   "RIO3 Tanks Pressure Switch Hi Hi" : Bool = PLC "RIO3 Tanks Pressure Switch Hi Hi" AT %I33.1, 1 s
   "RIO3_SPR_DI_27_6" : Bool = PLC RIO3_SPR_DI_27_6 AT %I27.6, 1 s
   "RIO3_SPR_DI_27_7" : Bool = PLC RIO3_SPR_DI_27_7 AT %I27.7, 1 s
   "RIO3_SPR_DI_30_6" : Bool = PLC RIO3_SPR_DI_30_6 AT %I30.6, 1 s
   "RIO3_SPR_DI_30_7" : Bool = PLC RIO3_SPR_DI_30_7 AT %I30.7, 1 s
   "RIO3_SPR_DI_33_3" : Bool = PLC RIO3_SPR_DI_33_3 AT %I33.3, 1 s
   "RIO3_SPR_DI_33_4" : Bool = PLC RIO3_SPR_DI_33_4 AT %I33.4, 1 s
   "RIO3_SPR_DI_33_5" : Bool = PLC RIO3_SPR_DI_33_5 AT %I33.5, 1 s
   "RIO3_SPR_DI_33_6" : Bool = PLC RIO3_SPR_DI_33_6 AT %I33.6, 1 s
   "RIO3_SPR_DI_33_7" : Bool = PLC RIO3_SPR_DI_33_7 AT %I33.7, 1 s
   "RIO4 Tanks Pressure Switch Hi Hi" : Bool = PLC "RIO4 Tanks Pressure Switch Hi Hi" AT %I45.1, 1 s
   "RIO4_SPR_DI_139_6" : Bool = PLC RIO4_SPR_DI_139_6 AT %I39.6, 1 s
   "RIO4_SPR_DI_139_7" : Bool = PLC RIO4_SPR_DI_139_7 AT %I39.7, 1 s
   "RIO4_SPR_DI_142_6" : Bool = PLC RIO4_SPR_DI_142_6 AT %I42.6, 1 s
   "RIO4_SPR_DI_142_7" : Bool = PLC RIO4_SPR_DI_142_7 AT %I42.7, 1 s
   "RIO4_SPR_DI_145_3" : Bool = PLC RIO4_SPR_DI_145_3 AT %I45.3, 1 s
   "RIO4_SPR_DI_145_4" : Bool = PLC RIO4_SPR_DI_145_4 AT %I45.4, 1 s
   "RIO4_SPR_DI_145_5" : Bool = PLC RIO4_SPR_DI_145_5 AT %I45.5, 1 s
   "RIO4_SPR_DI_145_6" : Bool = PLC RIO4_SPR_DI_145_6 AT %I45.6, 1 s
   "RIO4_SPR_DI_145_7" : Bool = PLC RIO4_SPR_DI_145_7 AT %I45.7, 1 s
   "RIO5 Tanks Pressure Switch Hi Hi" : Bool = PLC "RIO5 Tanks Pressure Switch Hi Hi" AT %I57.1, 1 s
   "RIO5_SPR_DI_51_6" : Bool = PLC RIO5_SPR_DI_51_6 AT %I51.6, 1 s
   "RIO5_SPR_DI_51_7" : Bool = PLC RIO5_SPR_DI_51_7 AT %I51.7, 1 s
   "RIO5_SPR_DI_54_6" : Bool = PLC RIO5_SPR_DI_54_6 AT %I54.6, 1 s
   "RIO5_SPR_DI_54_7" : Bool = PLC RIO5_SPR_DI_54_7 AT %I54.7, 1 s
   "RIO5_SPR_DI_57_3" : Bool = PLC RIO5_SPR_DI_57_3 AT %I57.3, 1 s
   "RIO5_SPR_DI_57_4" : Bool = PLC RIO5_SPR_DI_57_4 AT %I57.4, 1 s
   "RIO5_SPR_DI_57_5" : Bool = PLC RIO5_SPR_DI_57_5 AT %I57.5, 1 s
   "RIO5_SPR_DI_57_6" : Bool = PLC RIO5_SPR_DI_57_6 AT %I57.6, 1 s
   "RIO5_SPR_DI_57_7" : Bool = PLC RIO5_SPR_DI_57_7 AT %I57.7, 1 s
   "RIO6 Tanks Pressure Switch Hi Hi" : Bool = PLC "RIO6 Tanks Pressure Switch Hi Hi" AT %I66.1, 1 s
   "RIO6_SPR_DI_60_6" : Bool = PLC RIO6_SPR_DI_60_6 AT %I60.6, 1 s
   "RIO6_SPR_DI_60_7" : Bool = PLC RIO6_SPR_DI_60_7 AT %I60.7, 1 s
   "RIO6_SPR_DI_63_6" : Bool = PLC RIO6_SPR_DI_63_6 AT %I63.6, 1 s
   "RIO6_SPR_DI_63_7" : Bool = PLC RIO6_SPR_DI_63_7 AT %I63.7, 1 s
   "RIO6_SPR_DI_66_3" : Bool = PLC RIO6_SPR_DI_66_3 AT %I66.3, 1 s
   "RIO6_SPR_DI_66_4" : Bool = PLC RIO6_SPR_DI_66_4 AT %I66.4, 1 s
   "RIO6_SPR_DI_66_5" : Bool = PLC RIO6_SPR_DI_66_5 AT %I66.5, 1 s
   "RIO6_SPR_DI_66_6" : Bool = PLC RIO6_SPR_DI_66_6 AT %I66.6, 1 s
   "RIO6_SPR_DI_66_7" : Bool = PLC RIO6_SPR_DI_66_7 AT %I66.7, 1 s
   "RIO7 Tank Pressure Switch Hi Hi" : Bool = PLC "RIO7 Tank Pressure Switch Hi Hi" AT %I78.1, 1 s
   "RIO7_SPR_DI_175_6" : Bool = PLC RIO7_SPR_DI_175_6 AT %I75.6, 1 s
   "RIO7_SPR_DI_175_7" : Bool = PLC RIO7_SPR_DI_175_7 AT %I75.7, 1 s
   "RIO7_SPR_DI_178_2" : Bool = PLC RIO7_SPR_DI_178_2 AT %I78.2, 1 s
   "RIO7_SPR_DI_178_3" : Bool = PLC RIO7_SPR_DI_178_3 AT %I78.3, 1 s
   "RIO7_SPR_DI_178_4" : Bool = PLC RIO7_SPR_DI_178_4 AT %I78.4, 1 s
   "RIO7_SPR_DI_178_5" : Bool = PLC RIO7_SPR_DI_178_5 AT %I78.5, 1 s
   "RIO7_SPR_DI_178_6" : Bool = PLC RIO7_SPR_DI_178_6 AT %I78.6, 1 s
   "RIO7_SPR_DI_178_7" : Bool = PLC RIO7_SPR_DI_178_7 AT %I78.7, 1 s
   "Safety System Interlock" : Bool = PLC "10_DI_Data".SFTY_SYS_IL AT %DB1.DBX0.0, 1 s
   "Sequence Times_DB_De-Ox SP Time" : Real = PLC "Sequence Times_DB"."De-Ox SP Time", 1 s
   "Sequence Times_DB_De-Ox Time" : Real = PLC "Sequence Times_DB"."De-Ox Time", 1 s
   "Sequence Times_DB_De-Ox Timer_Days Left" : DInt = PLC "Sequence Times_DB"."De-Ox Timer"."Days Left", 1 s
   "Sequence Times_DB_De-Ox Timer_Hours Left" : DInt = PLC "Sequence Times_DB"."De-Ox Timer"."Hours Left", 1 s
   "Sequence Times_DB_De-Ox Timer_Minutes Left" : DInt = PLC "Sequence Times_DB"."De-Ox Timer"."Minutes Left", 1 s
   "Sequence Times_DB_De-Ox Timer_PT_HOURS" : Real = PLC "Sequence Times_DB"."De-Ox Timer".PT_HOURS, 1 s
   "Sequence Times_DB_Dwell" : Real = PLC "Sequence Times_DB"."Dwell Time", 1 s
   "Sequence Times_DB_Dwell Timer_Days Left" : DInt = PLC "Sequence Times_DB"."Dwell Timer"."Days Left", 1 s
   "Sequence Times_DB_Dwell Timer_Hours Left" : DInt = PLC "Sequence Times_DB"."Dwell Timer"."Hours Left", 1 s
   "Sequence Times_DB_Dwell Timer_Minutes Left" : DInt = PLC "Sequence Times_DB"."Dwell Timer"."Minutes Left", 1 s
   "Sequence Times_DB_Dwell Timer_PT_HOURS" : Real = PLC "Sequence Times_DB"."Dwell Timer".PT_HOURS, 1 s
   "Sequence Times_DB_Jurney Time" : Real = PLC "Sequence Times_DB"."Jurney Time", 1 s
   "Sequence Times_DB_Jurney Time FB_Days Left" : Int = PLC "Sequence Times_DB"."Jurney Time FB"."Days Left", 1 s
   "Sequence Times_DB_Jurney Time FB_Hours Left" : Int = PLC "Sequence Times_DB"."Jurney Time FB"."Hours Left", 1 s
   "Sequence Times_DB_Jurney Time FB_PT_DAYS" : Real = PLC "Sequence Times_DB"."Jurney Time FB".PT_DAYS, 1 s
   "Sequence Times_DB_Jurney Timer_PT_DAYS" : Real = PLC "Sequence Times_DB"."Jurney Timer".PT_DAYS, 1 s
   "Sequence Times_DB_Jurney Timer_PT_HOURS" : Real = PLC "Sequence Times_DB"."Jurney Timer".PT_HOURS, 1 s
   "Sequence Times_DB_Jurney Timer_PT_MINUTES" : Real = PLC "Sequence Times_DB"."Jurney Timer".PT_MINUTES, 1 s
   "Sequence Times_DB_Post-Dwell" : Real = PLC "Sequence Times_DB"."Post-Dwell Time", 1 s
   "Sequence Times_DB_Post-Dwell Remaining_Days Left" : DInt = PLC "Sequence Times_DB"."Post-Dwell Timer"."Days Left", 1 s
   "Sequence Times_DB_Post-Dwell Remaining_Hours Left" : DInt = PLC "Sequence Times_DB"."Post-Dwell Timer"."Hours Left", 1 s
   "Sequence Times_DB_Post-Dwell Remaining_Minutes Left" : DInt = PLC "Sequence Times_DB"."Post-Dwell Timer"."Minutes Left", 1 s
   "Sequence Times_DB_Post-Dwell Remaining_PT_HOURS" : Real = PLC "Sequence Times_DB"."Post-Dwell Timer".PT_HOURS, 1 s
   "Sequence Times_DB_Pre-Dwell Time" : Real = PLC "Sequence Times_DB"."Pre-Dwell Time", 1 s
   "Sequence Times_DB_Pre-Dwell Timer_Days Left" : DInt = PLC "Sequence Times_DB"."Pre-Dwell Timer"."Days Left", 1 s
   "Sequence Times_DB_Pre-Dwell Timer_Hours Left" : DInt = PLC "Sequence Times_DB"."Pre-Dwell Timer"."Hours Left", 1 s
   "Sequence Times_DB_Pre-Dwell Timer_Minutes Left" : DInt = PLC "Sequence Times_DB"."Pre-Dwell Timer"."Minutes Left", 1 s
   "Sequence Times_DB_Pre-Dwell Timer_PT_DAYS" : Real = PLC "Sequence Times_DB"."Pre-Dwell Timer".PT_DAYS, 1 s
   "Sequence Times_DB_Pre-Dwell Timer_PT_HOURS" : Real = PLC "Sequence Times_DB"."Pre-Dwell Timer".PT_HOURS, 1 s
   "Sequence Times_DB_Pre-Dwell Timer_PT_MINUTES" : Real = PLC "Sequence Times_DB"."Pre-Dwell Timer".PT_MINUTES, 1 s
   "Sequence Times_DB_Re-Ox Time" : Real = PLC "Sequence Times_DB"."Re-Ox Time", 1 s
   "Sequence Times_DB_Re-Ox Timer_Days Left" : DInt = PLC "Sequence Times_DB"."Re-Ox Timer"."Days Left", 1 s
   "Sequence Times_DB_Re-Ox Timer_Hours Left" : DInt = PLC "Sequence Times_DB"."Re-Ox Timer"."Hours Left", 1 s
   "Sequence Times_DB_Re-Ox Timer_Minutes Left" : DInt = PLC "Sequence Times_DB"."Re-Ox Timer"."Minutes Left", 1 s
   "Sequence Times_DB_Re-Ox Timer_PT_HOURS" : Real = PLC "Sequence Times_DB"."Re-Ox Timer".PT_HOURS, 1 s
   "Sequence Times_DB_Treatment Timer_Days" : DInt = PLC "Sequence Times_DB"."Treatment Timer".Days, 1 s
   "Sequence Times_DB_Treatment Timer_Days Left" : DInt = PLC "Sequence Times_DB"."Treatment Timer"."Days Left", 1 s
   "Sequence Times_DB_Treatment Timer_Enable" : Bool = PLC "Sequence Times_DB"."Treatment Timer".Enable, 1 s
   "Sequence Times_DB_Treatment Timer_Hours" : DInt = PLC "Sequence Times_DB"."Treatment Timer".Hours, 1 s
   "Sequence Times_DB_Treatment Timer_Hours Left" : DInt = PLC "Sequence Times_DB"."Treatment Timer"."Hours Left", 1 s
   "Sequence Times_DB_Treatment Timer_Minutes" : DInt = PLC "Sequence Times_DB"."Treatment Timer".Minutes, 1 s
   "Sequence Times_DB_Treatment Timer_Minutes Left" : DInt = PLC "Sequence Times_DB"."Treatment Timer"."Minutes Left", 1 s
   "Shell Cooling Water Level Hi Hi Switch" : Bool = PLC "10 DI_DATA".LS001 AT %DB1.DBX0.0, 1 s
   "Shell CSW Temp Scaled" : Real = PLC "12_AI_Data".TIT315_SCALED AT %DB1.DBX0.0, 1 s
   "Shutdown" : Bool = PLC "14_DQ_Data".24PF2 AT %DB1.DBX0.0, 1 s
   "Shutdown Alarm" : Bool = PLC "14_DQ_Data".24K3 AT %DB1.DBX0.0, 1 s
   "Silence Buzzer" : Bool = PLC "80_From_HMI".SLNCE_BZR AT %DB1.DBX0.0, 1 s
   "Soot System Opacity" : Bool = PLC "10 DI_DATA".E700_OPACITY AT %DB1.DBX0.0, 1 s
   "Soot System Power Healthy" : Bool = PLC "10 DI_DATA".E700_PWR_OK AT %DB1.DBX0.0, 1 s
   "Spare Output BC Q1.2" : Bool = PLC "14_DQ_Data".R2_SPR_DQ_1_2 AT %DB1.DBX0.0, 1 s
   "Spare Output BC Q1.3" : Bool = PLC "14_DQ_Data".R2_SPR_DQ_1_3 AT %DB1.DBX0.0, 1 s
   "Spare Output BC Q1.4" : Bool = PLC "14_DQ_Data".R2_SPR_DQ_1_4 AT %DB1.DBX0.0, 1 s
   "Spare Output BC Q1.5" : Bool = PLC "14_DQ_Data".R2_SPR_DQ_1_5 AT %DB1.DBX0.0, 1 s
   "Spare Output BC Q1.6" : Bool = PLC "14_DQ_Data".R2_SPR_DQ_1_6 AT %DB1.DBX0.0, 1 s
   "Spare Output IGG Q0.7" : Bool = PLC "14_DQ_Data".R2_SPR_DQ_0_7 AT %DB1.DBX0.0, 1 s
   "Spare Output IGG Q1.0" : Bool = PLC "14_DQ_Data".R2_SPR_DQ_1_0 AT %DB1.DBX0.0, 1 s
   "Start IGG Flag" : Bool = PLC "80_From_HMI".RUN_IGG AT %DB1.DBX0.0, 1 s
   "Start Sequenc_DB_Post Purge Time Sec" : Int, internal
   "Tank 1P BWT Level High High Switch" : Bool = PLC "Tank 1P BWT Level High High Switch" AT %I9.2, 1 s
   "Tank 1P GTT Isolation Valve Feedback - Closed" : Bool = PLC "Tank 1P GTT Isolation Valve Feedback - Closed" AT %I3.1, 1 s
   "Tank 1P GTT Isolation Valve Feedback - Opened" : Bool = PLC "Tank 1P GTT Isolation Valve Feedback - Opened" AT %I3.0, 1 s
   "Tank 1P Tank Vent Valve 1 Feedback - Closed" : Bool = PLC "Tank 1P Tank Vent Valve 1 Feedback - Closed" AT %I3.3, 1 s
   "Tank 1P Tank Vent Valve 1 Feedback - Opened" : Bool = PLC "Tank 1P Tank Vent Valve 1 Feedback - Opened" AT %I3.2, 1 s
   "Tank 1P Tank Vent Valve 2 Feedback - Closed" : Bool = PLC "Tank 1P Tank Vent Valve 2 Feedback - Closed" AT %I3.5, 1 s
   "Tank 1P Tank Vent Valve 2 Feedback - Opened" : Bool = PLC "Tank 1P Tank Vent Valve 2 Feedback - Opened" AT %I3.4, 1 s
   "Tank 1S BWT Level High High Switch" : Bool = PLC "Tank 1S BWT Level High High Switch" AT %I9.3, 1 s
   "Tank 1S GTT Isolation Valve Feedback - Closed" : Bool = PLC "Tank 1S GTT Isolation Valve Feedback - Closed" AT %I6.1, 1 s
   "Tank 1S GTT Isolation Valve Feedback - Opened" : Bool = PLC "Tank 1S GTT Isolation Valve Feedback - Opened" AT %I6.0, 1 s
   "Tank 1S Tank Vent Valve 1 Feedback - Closed" : Bool = PLC "Tank 1S Tank Vent Valve 1 Feedback - Closed" AT %I6.3, 1 s
   "Tank 1S Tank Vent Valve 1 Feedback - Opened" : Bool = PLC "Tank 1S Tank Vent Valve 1 Feedback - Opened" AT %I6.2, 1 s
   "Tank 1S Tank Vent Valve 2 Feedback - Closed" : Bool = PLC "Tank 1S Tank Vent Valve 2 Feedback - Closed" AT %I6.5, 1 s
   "Tank 1S Tank Vent Valve 2 Feedback - Opened" : Bool = PLC "Tank 1S Tank Vent Valve 2 Feedback - Opened" AT %I6.4, 1 s
   "Tank 2P BWT Level High High Switch" : Bool = PLC "Tank 2P BWT Level High High Switch" AT %I21.0, 1 s
   "Tank 2P GTT Isolation Valve Feedback - Closed" : Bool = PLC "Tank 2P GTT Isolation Valve Feedback - Closed" AT %I15.1, 1 s
   "Tank 2P GTT Isolation Valve Feedback - Opened" : Bool = PLC "Tank 2P GTT Isolation Valve Feedback - Opened" AT %I15.0, 1 s
   "Tank 2P Tank Vent Valve 1 Feedback - Closed" : Bool = PLC "Tank 2P Tank Vent Valve 1 Feedback - Closed" AT %I15.3, 1 s
   "Tank 2P Tank Vent Valve 1 Feedback - Opened" : Bool = PLC "Tank 2P Tank Vent Valve 1 Feedback - Opened" AT %I15.2, 1 s
   "Tank 2P Tank Vent Valve 2 Feedback - Closed" : Bool = PLC "Tank 2P Tank Vent Valve 2 Feedback - Closed" AT %I15.5, 1 s
   "Tank 2P Tank Vent Valve 2 Feedback - Opened" : Bool = PLC "Tank 2P Tank Vent Valve 2 Feedback - Opened" AT %I15.4, 1 s
   "Tank 2S BWT Level High High Switch" : Bool = PLC "Tank 2S BWT Level High High Switch" AT %I21.2, 1 s
   "Tank 2S GTT Isolation Valve Feedback - Closed" : Bool = PLC "Tank 2S GTT Isolation Valve Feedback - Closed" AT %I18.1, 1 s
   "Tank 2S GTT Isolation Valve Feedback - Opened" : Bool = PLC "Tank 2S GTT Isolation Valve Feedback - Opened" AT %I18.0, 1 s
   "Tank 2S Tank Vent Valve 1 Feedback - Closed" : Bool = PLC "Tank 2S Tank Vent Valve 1 Feedback - Closed" AT %I18.3, 1 s
   "Tank 2S Tank Vent Valve 1 Feedback - Opened" : Bool = PLC "Tank 2S Tank Vent Valve 1 Feedback - Opened" AT %I18.2, 1 s
   "Tank 2S Tank Vent Valve 2 Feedback - Closed" : Bool = PLC "Tank 2S Tank Vent Valve 2 Feedback - Closed" AT %I18.5, 1 s
   "Tank 2S Tank Vent Valve 2 Feedback - Opened" : Bool = PLC "Tank 2S Tank Vent Valve 2 Feedback - Opened" AT %I18.4, 1 s
   "Tank 3P BWT Level High High Switch" : Bool = PLC "Tank 3P BWT Level High High Switch" AT %I33.0, 1 s
   "Tank 3P GTT Isolation Valve Feedback - Closed" : Bool = PLC "Tank 3P GTT Isolation Valve Feedback - Closed" AT %I27.1, 1 s
   "Tank 3P GTT Isolation Valve Feedback - Opened" : Bool = PLC "Tank 3P GTT Isolation Valve Feedback - Opened" AT %I27.0, 1 s
   "Tank 3P Tank Vent Valve 1 Feedback - Closed" : Bool = PLC "Tank 3P Tank Vent Valve 1 Feedback - Closed" AT %I27.3, 1 s
   "Tank 3P Tank Vent Valve 1 Feedback - Opened" : Bool = PLC "Tank 3P Tank Vent Valve 1 Feedback - Opened" AT %I27.2, 1 s
   "Tank 3P Tank Vent Valve 2 Feedback - Closed" : Bool = PLC "Tank 3P Tank Vent Valve 2 Feedback - Closed" AT %I27.5, 1 s
   "Tank 3P Tank Vent Valve 2 Feedback - Opened" : Bool = PLC "Tank 3P Tank Vent Valve 2 Feedback - Opened" AT %I27.4, 1 s
   "Tank 3S BWT Level High High Switch" : Bool = PLC "Tank 3S BWT Level High High Switch" AT %I33.2, 1 s
   "Tank 3S GTT Isolation Valve Feedback - Closed" : Bool = PLC "Tank 3S GTT Isolation Valve Feedback - Closed" AT %I30.1, 1 s
   "Tank 3S GTT Isolation Valve Feedback - Opened" : Bool = PLC "Tank 3S GTT Isolation Valve Feedback - Opened" AT %I30.0, 1 s
   "Tank 3S Tank Vent Valve 1 Feedback - Closed" : Bool = PLC "Tank 3S Tank Vent Valve 1 Feedback - Closed" AT %I30.3, 1 s
   "Tank 3S Tank Vent Valve 1 Feedback - Opened" : Bool = PLC "Tank 3S Tank Vent Valve 1 Feedback - Opened" AT %I30.2, 1 s
   "Tank 3S Tank Vent Valve 2 Feedback - Closed" : Bool = PLC "Tank 3S Tank Vent Valve 2 Feedback - Closed" AT %I30.5, 1 s
   "Tank 3S Tank Vent Valve 2 Feedback - Opened" : Bool = PLC "Tank 3S Tank Vent Valve 2 Feedback - Opened" AT %I30.4, 1 s
   "Tank 4P BWT Level High High Switch" : Bool = PLC "Tank 4P BWT Level High High Switch" AT %I45.0, 1 s
   "Tank 4P GTT Isolation Valve Feedback - Closed" : Bool = PLC "Tank 4P GTT Isolation Valve Feedback - Closed" AT %I39.1, 1 s
   "Tank 4P GTT Isolation Valve Feedback - Opened" : Bool = PLC "Tank 4P GTT Isolation Valve Feedback - Opened" AT %I39.0, 1 s
   "Tank 4P Tank Vent Valve 1 Feedback - Closed" : Bool = PLC "Tank 4P Tank Vent Valve 1 Feedback - Closed" AT %I39.3, 1 s
   "Tank 4P Tank Vent Valve 1 Feedback - Opened" : Bool = PLC "Tank 4P Tank Vent Valve 1 Feedback - Opened" AT %I39.2, 1 s
   "Tank 4P Tank Vent Valve 2 Feedback - Closed" : Bool = PLC "Tank 4P Tank Vent Valve 2 Feedback - Closed" AT %I39.5, 1 s
   "Tank 4P Tank Vent Valve 2 Feedback - Opened" : Bool = PLC "Tank 4P Tank Vent Valve 2 Feedback - Opened" AT %I39.4, 1 s
   "Tank 4S BWT Level High High Switch" : Bool = PLC "Tank 4S BWT Level High High Switch" AT %I45.2, 1 s
   "Tank 4S GTT Isolation Valve Feedback - Closed" : Bool = PLC "Tank 4S GTT Isolation Valve Feedback - Closed" AT %I42.1, 1 s
   "Tank 4S GTT Isolation Valve Feedback - Opened" : Bool = PLC "Tank 4S GTT Isolation Valve Feedback - Opened" AT %I42.0, 1 s
   "Tank 4S Tank Vent Valve 1 Feedback - Closed" : Bool = PLC "Tank 4S Tank Vent Valve 1 Feedback - Closed" AT %I42.3, 1 s
   "Tank 4S Tank Vent Valve 1 Feedback - Opened" : Bool = PLC "Tank 4S Tank Vent Valve 1 Feedback - Opened" AT %I42.2, 1 s
   "Tank 4S Tank Vent Valve 2 Feedback - Closed" : Bool = PLC "Tank 4S Tank Vent Valve 2 Feedback - Closed" AT %I42.5, 1 s
   "Tank 4S Tank Vent Valve 2 Feedback - Opened" : Bool = PLC "Tank 4S Tank Vent Valve 2 Feedback - Opened" AT %I42.4, 1 s
   "Tank 5P BWT Level High High Switch" : Bool = PLC "Tank 5P BWT Level High High Switch" AT %I57.0, 1 s
   "Tank 5P GTT Isolation Valve Feedback - Closed" : Bool = PLC "Tank 5P GTT Isolation Valve Feedback - Closed" AT %I51.1, 1 s
   "Tank 5P GTT Isolation Valve Feedback - Opened" : Bool = PLC "Tank 5P GTT Isolation Valve Feedback - Opened" AT %I51.0, 1 s
   "Tank 5P Tank Vent Valve 1 Feedback - Closed" : Bool = PLC "Tank 5P Tank Vent Valve 1 Feedback - Closed" AT %I51.3, 1 s
   "Tank 5P Tank Vent Valve 1 Feedback - Opened" : Bool = PLC "Tank 5P Tank Vent Valve 1 Feedback - Opened" AT %I51.2, 1 s
   "Tank 5P Tank Vent Valve 2 Feedback - Closed" : Bool = PLC "Tank 5P Tank Vent Valve 2 Feedback - Closed" AT %I51.5, 1 s
   "Tank 5P Tank Vent Valve 2 Feedback - Opened" : Bool = PLC "Tank 5P Tank Vent Valve 2 Feedback - Opened" AT %I51.4, 1 s
   "Tank 5S BWT Level High High Switch" : Bool = PLC "Tank 5S BWT Level High High Switch" AT %I57.2, 1 s
   "Tank 6P BWT Level High High Switch" : Bool = PLC "Tank 6P BWT Level High High Switch" AT %I66.0, 1 s
   "Tank 6S BWT Level High High Switch" : Bool = PLC "Tank 6S BWT Level High High Switch" AT %I66.2, 1 s
   "Test Pressure Valve Control" : Bool = PLC "14_DQ_Data".200CV127ControlOut AT %DB1.DBX0.0, 1 s
   "TIT406_ALM_ANALOG_DB74_HIGH LEVEL VALUE (H)" : Real = PLC TIT406_ALM_ANALOG_DB74."HIGH LEVEL VALUE (H)" AT %DB74.DBD30, 1 s
   "TIT406_ALM_ANALOG_DB74_LOW LEVEL VALUE (L)" : Real = PLC TIT406_ALM_ANALOG_DB74."LOW LEVEL VALUE (L)" AT %DB74.DBD26, 1 s
   "TIT406_ALM_ANALOG_DB74_VERY HIGH LEVEL VALUE (HH)" : Real = PLC TIT406_ALM_ANALOG_DB74."VERY HIGH LEVEL VALUE (HH)" AT %DB74.DBD34, 1 s
   "TIT406_ALM_ANALOG_DB74_VERY LOW LEVEL VALUE (LL)" : Real = PLC TIT406_ALM_ANALOG_DB74."VERY LOW LEVEL VALUE (LL)" AT %DB74.DBD22, 1 s
   "TIT408_ALM_ANALOG_DB75_HIGH LEVEL VALUE (H)" : Real = PLC TIT408_ALM_ANALOG_DB75."HIGH LEVEL VALUE (H)" AT %DB75.DBD30, 1 s
   "TIT408_ALM_ANALOG_DB75_LOW LEVEL VALUE (L)" : Real = PLC TIT408_ALM_ANALOG_DB75."LOW LEVEL VALUE (L)" AT %DB75.DBD26, 1 s
   "TIT408_ALM_ANALOG_DB75_VERY HIGH LEVEL VALUE (HH)" : Real = PLC TIT408_ALM_ANALOG_DB75."VERY HIGH LEVEL VALUE (HH)" AT %DB75.DBD34, 1 s
   "TIT408_ALM_ANALOG_DB75_VERY LOW LEVEL VALUE (LL)" : Real = PLC TIT408_ALM_ANALOG_DB75."VERY LOW LEVEL VALUE (LL)" AT %DB75.DBD22, 1 s
   "Treatment Runs Completed" : Bool = PLC "2102_TIME_CALCS_DB".POST_DWELL_TMR_DN AT %DB1.DBD0, 1 s
   "user_group" : Int, internal
   "Vent Valve Control HMI Position" : Real = PLC "16_AQ_Data".CV403_CNTRL AT %DB1.DBX0.0, 1 s
   "Vent Valve Position Control" : Real = PLC "12_AI_Data".CV403_SCALED AT %DB1.DBX0.0, 1 s
   "Voyage_TIME_exceded" : Bool = PLC "2102_TIME_CALCS_DB".Voyage_TIME_invalid AT %DB1.DBW0, 1 s
   "Warning Alarm" : Bool = PLC "14_DQ_Data".24PF3 AT %DB1.DBX0.0, 1 s
   "Sequence Times_DB_Continue" : Bool = PLC "Sequence Times_DB".Continue, 1 s
   "Recipe Tag" : Int AT %DB1.DBX0.0
   "Record Data Tag" : Int AT %DB1.DBX0.0
   "Data_From_WBT_Level_APT" : Real = PLC Data_From_WBT.Level_APT, 1 s
   "Data_From_WBT_Level_WBT_6P" : Real = PLC Data_From_WBT.Level_WBT_6P, 1 s
   "Data_From_WBT_Level_WBT_5P" : Real = PLC Data_From_WBT.Level_WBT_5P, 1 s
   "Data_From_WBT_Level_WBT_4P" : Real = PLC Data_From_WBT.Level_WBT_4P, 1 s
   "Data_From_WBT_Level_WBT_3P" : Real = PLC Data_From_WBT.Level_WBT_3P, 1 s
   "Data_From_WBT_Level_WBT_2P" : Real = PLC Data_From_WBT.Level_WBT_2P, 1 s
   "Data_From_WBT_Level_WBT_1P" : Real = PLC Data_From_WBT.Level_WBT_1P, 1 s
   "Data_From_WBT_Level_FPT" : Real = PLC Data_From_WBT.Level_FPT, 1 s
   "Data_From_WBT_Level_WBT_1S" : Real = PLC Data_From_WBT.Level_WBT_1S, 1 s
   "Data_From_WBT_Level_WBT_2S" : Real = PLC Data_From_WBT.Level_WBT_2S, 1 s
   "Data_From_WBT_Level_WBT_3S" : Real = PLC Data_From_WBT.Level_WBT_3S, 1 s
   "Data_From_WBT_Level_WBT_4S" : Real = PLC Data_From_WBT.Level_WBT_4S, 1 s
   "Data_From_WBT_Level_WBT_5S" : Real = PLC Data_From_WBT.Level_WBT_5S, 1 s
   "Data_From_WBT_Level_WBT_6S" : Real = PLC Data_From_WBT.Level_WBT_6S, 1 s
   "IN_Level_APT" : Int = PLC IN_Level_APT AT %IW1026, 1 s
   "Data_From_WBT_Level_APT m" : Real = PLC Data_From_WBT."Level_APT m", 1 s
   "Data_From_WBT_Level_WBT_6S m" : Real = PLC Data_From_WBT."Level_WBT_6S m", 1 s
   "Data_From_WBT_Level_WBT_5S m" : Real = PLC Data_From_WBT."Level_WBT_5S m", 1 s
   "Data_From_WBT_Level_WBT_4S m" : Real = PLC Data_From_WBT."Level_WBT_4S m", 1 s
   "Data_From_WBT_Level_WBT_3S m" : Real = PLC Data_From_WBT."Level_WBT_3S m", 1 s
   "Data_From_WBT_Level_WBT_2S m" : Real = PLC Data_From_WBT."Level_WBT_2S m", 1 s
   "Data_From_WBT_Level_WBT_1S m" : Real = PLC Data_From_WBT."Level_WBT_1S m", 1 s
   "Data_From_WBT_Level_FPT m" : Real = PLC Data_From_WBT."Level_FPT m", 1 s
   "Data_From_WBT_Level_WBT_1P m" : Real = PLC Data_From_WBT."Level_WBT_1P m", 1 s
   "Data_From_WBT_Level_WBT_2P m" : Real = PLC Data_From_WBT."Level_WBT_2P m", 1 s
   "Data_From_WBT_Level_WBT_3P m" : Real = PLC Data_From_WBT."Level_WBT_3P m", 1 s
   "Data_From_WBT_Level_WBT_4P m" : Real = PLC Data_From_WBT."Level_WBT_4P m", 1 s
   "Data_From_WBT_Level_WBT_5P m" : Real = PLC Data_From_WBT."Level_WBT_5P m", 1 s
   "Data_From_WBT_Level_WBT_6P m" : Real = PLC Data_From_WBT."Level_WBT_6P m", 1 s
   "Alarm beacon handling_DB_Warning" : Bool = PLC "Alarm beacon handling_DB".Warning, 1 s
   "Alarm beacon handling_DB_Alarm" : Bool = PLC "Alarm beacon handling_DB".Alarm, 1 s
   "63_Safety System Interlock_IDB_Lockout Healthy" : Bool = PLC "63_Safety System Interlock_IDB"."Lockout Healthy", 1 s
   "63_Safety System Interlock_IDB_Reset Lockout" : Bool = PLC "63_Safety System Interlock_IDB"."Reset Lockout", 1 s
   "IDB_E131_Functioning Hours_Service Time bit" : Bool = PLC "IDB_E131_Functioning Hours"."Service Time bit", 1 s
   "Operation hours E139_IDB_Service Time bit" : Bool = PLC "Operation hours E139_IDB"."Service Time bit", 1 s
   "E-400 Animation_DB_Animation" : Int = PLC "E-400 Animation_DB".Animation, 1 s
   "20_TANKS_IP_DATA_RIO_01_FIRST_TANK_TANK_ALARM" : Bool = PLC "20_TANKS_IP_DATA".RIO_01.FIRST_TANK.TANK_ALARM, 1 s
   "CSW_Animation_DB_Animation" : Int = PLC CSW_Animation_DB.Animation, 1 s
   "103_Main_Burner_DB_FLM_DET" : Bool = PLC "103_Main_Burner_DB".FLM_DET, 1 s
   "504_Tank Grouping_DB2020_Time Left Tank_Time Left d Tank 1" : DInt = PLC "504_Tank Grouping_DB2020"."Time Left Tank"."Time Left d Tank 1", 1 s
   "504_Tank Grouping_DB2020_Time Left Tank_Time Left d Tank 10" : DInt = PLC "504_Tank Grouping_DB2020"."Time Left Tank"."Time Left d Tank 10", 1 s
   "504_Tank Grouping_DB2020_Time Left Tank_Time Left d Tank 11" : DInt = PLC "504_Tank Grouping_DB2020"."Time Left Tank"."Time Left d Tank 11", 1 s
   "504_Tank Grouping_DB2020_Time Left Tank_Time Left d Tank 12" : DInt = PLC "504_Tank Grouping_DB2020"."Time Left Tank"."Time Left d Tank 12", 1 s
   "504_Tank Grouping_DB2020_Time Left Tank_Time Left d Tank 13" : DInt = PLC "504_Tank Grouping_DB2020"."Time Left Tank"."Time Left d Tank 13", 1 s
   "504_Tank Grouping_DB2020_Time Left Tank_Time Left d Tank 14" : DInt = PLC "504_Tank Grouping_DB2020"."Time Left Tank"."Time Left d Tank 14", 1 s
   "504_Tank Grouping_DB2020_Time Left Tank_Time Left d Tank 2" : DInt = PLC "504_Tank Grouping_DB2020"."Time Left Tank"."Time Left d Tank 2", 1 s
   "504_Tank Grouping_DB2020_Time Left Tank_Time Left d Tank 3" : DInt = PLC "504_Tank Grouping_DB2020"."Time Left Tank"."Time Left d Tank 3", 1 s
   "504_Tank Grouping_DB2020_Time Left Tank_Time Left d Tank 4" : DInt = PLC "504_Tank Grouping_DB2020"."Time Left Tank"."Time Left d Tank 4", 1 s
   "504_Tank Grouping_DB2020_Time Left Tank_Time Left d Tank 5" : DInt = PLC "504_Tank Grouping_DB2020"."Time Left Tank"."Time Left d Tank 5", 1 s
   "504_Tank Grouping_DB2020_Time Left Tank_Time Left d Tank 6" : DInt = PLC "504_Tank Grouping_DB2020"."Time Left Tank"."Time Left d Tank 6", 1 s
   "504_Tank Grouping_DB2020_Time Left Tank_Time Left d Tank 7" : DInt = PLC "504_Tank Grouping_DB2020"."Time Left Tank"."Time Left d Tank 7", 1 s
   "504_Tank Grouping_DB2020_Time Left Tank_Time Left d Tank 8" : DInt = PLC "504_Tank Grouping_DB2020"."Time Left Tank"."Time Left d Tank 8", 1 s
   "504_Tank Grouping_DB2020_Time Left Tank_Time Left d Tank 9" : DInt = PLC "504_Tank Grouping_DB2020"."Time Left Tank"."Time Left d Tank 9", 1 s
   "504_Tank Grouping_DB2020_Time Left Tank_Time Left h Tank 1" : DInt = PLC "504_Tank Grouping_DB2020"."Time Left Tank"."Time Left h Tank 1", 1 s
   "504_Tank Grouping_DB2020_Time Left Tank_Time Left h Tank 10" : DInt = PLC "504_Tank Grouping_DB2020"."Time Left Tank"."Time Left h Tank 10", 1 s
   "504_Tank Grouping_DB2020_Time Left Tank_Time Left h Tank 11" : DInt = PLC "504_Tank Grouping_DB2020"."Time Left Tank"."Time Left h Tank 11", 1 s
   "504_Tank Grouping_DB2020_Time Left Tank_Time Left h Tank 12" : DInt = PLC "504_Tank Grouping_DB2020"."Time Left Tank"."Time Left h Tank 12", 1 s
   "504_Tank Grouping_DB2020_Time Left Tank_Time Left h Tank 13" : DInt = PLC "504_Tank Grouping_DB2020"."Time Left Tank"."Time Left h Tank 13", 1 s
   "504_Tank Grouping_DB2020_Time Left Tank_Time Left h Tank 14" : DInt = PLC "504_Tank Grouping_DB2020"."Time Left Tank"."Time Left h Tank 14", 1 s
   "504_Tank Grouping_DB2020_Time Left Tank_Time Left h Tank 2" : DInt = PLC "504_Tank Grouping_DB2020"."Time Left Tank"."Time Left h Tank 2", 1 s
   "504_Tank Grouping_DB2020_Time Left Tank_Time Left h Tank 3" : DInt = PLC "504_Tank Grouping_DB2020"."Time Left Tank"."Time Left h Tank 3", 1 s
   "504_Tank Grouping_DB2020_Time Left Tank_Time Left h Tank 4" : DInt = PLC "504_Tank Grouping_DB2020"."Time Left Tank"."Time Left h Tank 4", 1 s
   "504_Tank Grouping_DB2020_Time Left Tank_Time Left h Tank 5" : DInt = PLC "504_Tank Grouping_DB2020"."Time Left Tank"."Time Left h Tank 5", 1 s
   "504_Tank Grouping_DB2020_Time Left Tank_Time Left h Tank 6" : DInt = PLC "504_Tank Grouping_DB2020"."Time Left Tank"."Time Left h Tank 6", 1 s
   "504_Tank Grouping_DB2020_Time Left Tank_Time Left h Tank 7" : DInt = PLC "504_Tank Grouping_DB2020"."Time Left Tank"."Time Left h Tank 7", 1 s
   "504_Tank Grouping_DB2020_Time Left Tank_Time Left h Tank 8" : DInt = PLC "504_Tank Grouping_DB2020"."Time Left Tank"."Time Left h Tank 8", 1 s
   "504_Tank Grouping_DB2020_Time Left Tank_Time Left h Tank 9" : DInt = PLC "504_Tank Grouping_DB2020"."Time Left Tank"."Time Left h Tank 9", 1 s
   "504_Tank Grouping_DB2020_Time Left Tank_Time Left m Tank 1" : DInt = PLC "504_Tank Grouping_DB2020"."Time Left Tank"."Time Left m Tank 1", 1 s
   "504_Tank Grouping_DB2020_Time Left Tank_Time Left m Tank 10" : DInt = PLC "504_Tank Grouping_DB2020"."Time Left Tank"."Time Left m Tank 10", 1 s
   "504_Tank Grouping_DB2020_Time Left Tank_Time Left m Tank 11" : DInt = PLC "504_Tank Grouping_DB2020"."Time Left Tank"."Time Left m Tank 11", 1 s
   "504_Tank Grouping_DB2020_Time Left Tank_Time Left m Tank 12" : DInt = PLC "504_Tank Grouping_DB2020"."Time Left Tank"."Time Left m Tank 12", 1 s
   "504_Tank Grouping_DB2020_Time Left Tank_Time Left m Tank 13" : DInt = PLC "504_Tank Grouping_DB2020"."Time Left Tank"."Time Left m Tank 13", 1 s
   "504_Tank Grouping_DB2020_Time Left Tank_Time Left m Tank 14" : DInt = PLC "504_Tank Grouping_DB2020"."Time Left Tank"."Time Left m Tank 14", 1 s
   "504_Tank Grouping_DB2020_Time Left Tank_Time Left m Tank 2" : DInt = PLC "504_Tank Grouping_DB2020"."Time Left Tank"."Time Left m Tank 2", 1 s
   "504_Tank Grouping_DB2020_Time Left Tank_Time Left m Tank 3" : DInt = PLC "504_Tank Grouping_DB2020"."Time Left Tank"."Time Left m Tank 3", 1 s
   "504_Tank Grouping_DB2020_Time Left Tank_Time Left m Tank 4" : DInt = PLC "504_Tank Grouping_DB2020"."Time Left Tank"."Time Left m Tank 4", 1 s
   "504_Tank Grouping_DB2020_Time Left Tank_Time Left m Tank 5" : DInt = PLC "504_Tank Grouping_DB2020"."Time Left Tank"."Time Left m Tank 5", 1 s
   "504_Tank Grouping_DB2020_Time Left Tank_Time Left m Tank 6" : DInt = PLC "504_Tank Grouping_DB2020"."Time Left Tank"."Time Left m Tank 6", 1 s
   "504_Tank Grouping_DB2020_Time Left Tank_Time Left m Tank 7" : DInt = PLC "504_Tank Grouping_DB2020"."Time Left Tank"."Time Left m Tank 7", 1 s
   "504_Tank Grouping_DB2020_Time Left Tank_Time Left m Tank 8" : DInt = PLC "504_Tank Grouping_DB2020"."Time Left Tank"."Time Left m Tank 8", 1 s
   "504_Tank Grouping_DB2020_Time Left Tank_Time Left m Tank 9" : DInt = PLC "504_Tank Grouping_DB2020"."Time Left Tank"."Time Left m Tank 9", 1 s
   "TT002_ALM_ANALOG_DB76_HIGH LEVEL VALUE (H)" : Real = PLC TT002_ALM_ANALOG_DB76."HIGH LEVEL VALUE (H)" AT %DB76.DBD30, 1 s
   "TT002_ALM_ANALOG_DB76_LOW LEVEL VALUE (L)" : Real = PLC TT002_ALM_ANALOG_DB76."LOW LEVEL VALUE (L)" AT %DB76.DBD26, 1 s
   "TT002_ALM_ANALOG_DB76_VERY HIGH LEVEL VALUE (HH)" : Real = PLC TT002_ALM_ANALOG_DB76."VERY HIGH LEVEL VALUE (HH)" AT %DB76.DBD34, 1 s
   "TT002_ALM_ANALOG_DB76_VERY LOW LEVEL VALUE (LL)" : Real = PLC TT002_ALM_ANALOG_DB76."VERY LOW LEVEL VALUE (LL)" AT %DB76.DBD22, 1 s
   "TT426_1P_ALM_ANALOG_DB_HIGH LEVEL VALUE (H)" : Real = PLC TT426_1P_ALM_ANALOG_DB."HIGH LEVEL VALUE (H)" AT %DB2075.DBD30, 1 s
   "TT426_1P_ALM_ANALOG_DB_LOW LEVEL VALUE (L)" : Real = PLC TT426_1P_ALM_ANALOG_DB."LOW LEVEL VALUE (L)" AT %DB2075.DBD26, 1 s
   "TT426_1P_ALM_ANALOG_DB_VERY HIGH LEVEL VALUE (HH)" : Real = PLC TT426_1P_ALM_ANALOG_DB."VERY HIGH LEVEL VALUE (HH)" AT %DB2075.DBD34, 1 s
   "TT426_1P_ALM_ANALOG_DB_VERY LOW LEVEL VALUE (LL)" : Real = PLC TT426_1P_ALM_ANALOG_DB."VERY LOW LEVEL VALUE (LL)" AT %DB2075.DBD22, 1 s
   "TT426_1S_ALM_ANALOG_DB_HIGH LEVEL VALUE (H)" : Real = PLC TT426_1S_ALM_ANALOG_DB."HIGH LEVEL VALUE (H)" AT %DB2076.DBD30, 1 s
   "TT426_1S_ALM_ANALOG_DB_LOW LEVEL VALUE (L)" : Real = PLC TT426_1S_ALM_ANALOG_DB."LOW LEVEL VALUE (L)" AT %DB2076.DBD26, 1 s
   "TT426_1S_ALM_ANALOG_DB_VERY HIGH LEVEL VALUE (HH)" : Real = PLC TT426_1S_ALM_ANALOG_DB."VERY HIGH LEVEL VALUE (HH)" AT %DB2076.DBD34, 1 s
   "TT426_1S_ALM_ANALOG_DB_VERY LOW LEVEL VALUE (LL)" : Real = PLC TT426_1S_ALM_ANALOG_DB."VERY LOW LEVEL VALUE (LL)" AT %DB2076.DBD22, 1 s
   "TT426_3P_ALM_ANALOG_DB_HIGH LEVEL VALUE (H)" : Real = PLC TT426_3P_ALM_ANALOG_DB."HIGH LEVEL VALUE (H)" AT %DB2077.DBD30, 1 s
   "TT426_3P_ALM_ANALOG_DB_LOW LEVEL VALUE (L)" : Real = PLC TT426_3P_ALM_ANALOG_DB."LOW LEVEL VALUE (L)" AT %DB2077.DBD26, 1 s
   "TT426_3P_ALM_ANALOG_DB_VERY HIGH LEVEL VALUE (HH)" : Real = PLC TT426_3P_ALM_ANALOG_DB."VERY HIGH LEVEL VALUE (HH)" AT %DB2077.DBD34, 1 s
   "TT426_3P_ALM_ANALOG_DB_VERY LOW LEVEL VALUE (LL)" : Real = PLC TT426_3P_ALM_ANALOG_DB."VERY LOW LEVEL VALUE (LL)" AT %DB2077.DBD22, 1 s
   "TT426_3S_ALM_ANALOG_DB_HIGH LEVEL VALUE (H)" : Real = PLC TT426_3S_ALM_ANALOG_DB."HIGH LEVEL VALUE (H)" AT %DB2078.DBD30, 1 s
   "TT426_3S_ALM_ANALOG_DB_LOW LEVEL VALUE (L)" : Real = PLC TT426_3S_ALM_ANALOG_DB."LOW LEVEL VALUE (L)" AT %DB2078.DBD26, 1 s
   "TT426_3S_ALM_ANALOG_DB_VERY HIGH LEVEL VALUE (HH)" : Real = PLC TT426_3S_ALM_ANALOG_DB."VERY HIGH LEVEL VALUE (HH)" AT %DB2078.DBD34, 1 s
   "TT426_3S_ALM_ANALOG_DB_VERY LOW LEVEL VALUE (LL)" : Real = PLC TT426_3S_ALM_ANALOG_DB."VERY LOW LEVEL VALUE (LL)" AT %DB2078.DBD22, 1 s
   "TT426_4P_ALM_ANALOG_DB_HIGH LEVEL VALUE (H)" : Real = PLC TT426_4P_ALM_ANALOG_DB."HIGH LEVEL VALUE (H)" AT %DB2079.DBD30, 1 s
   "TT426_4P_ALM_ANALOG_DB_LOW LEVEL VALUE (L)" : Real = PLC TT426_4P_ALM_ANALOG_DB."LOW LEVEL VALUE (L)" AT %DB2079.DBD26, 1 s
   "TT426_4P_ALM_ANALOG_DB_VERY HIGH LEVEL VALUE (HH)" : Real = PLC TT426_4P_ALM_ANALOG_DB."VERY HIGH LEVEL VALUE (HH)" AT %DB2079.DBD34, 1 s
   "TT426_4P_ALM_ANALOG_DB_VERY LOW LEVEL VALUE (LL)" : Real = PLC TT426_4P_ALM_ANALOG_DB."VERY LOW LEVEL VALUE (LL)" AT %DB2079.DBD22, 1 s
   "TT426_4S_ALM_ANALOG_DB_HIGH LEVEL VALUE (H)" : Real = PLC TT426_4S_ALM_ANALOG_DB."HIGH LEVEL VALUE (H)" AT %DB2080.DBD30, 1 s
   "TT426_4S_ALM_ANALOG_DB_LOW LEVEL VALUE (L)" : Real = PLC TT426_4S_ALM_ANALOG_DB."LOW LEVEL VALUE (L)" AT %DB2080.DBD26, 1 s
   "TT426_4S_ALM_ANALOG_DB_VERY HIGH LEVEL VALUE (HH)" : Real = PLC TT426_4S_ALM_ANALOG_DB."VERY HIGH LEVEL VALUE (HH)" AT %DB2080.DBD34, 1 s
   "TT426_4S_ALM_ANALOG_DB_VERY LOW LEVEL VALUE (LL)" : Real = PLC TT426_4S_ALM_ANALOG_DB."VERY LOW LEVEL VALUE (LL)" AT %DB2080.DBD22, 1 s
   "TT426_5P_ALM_ANALOG_DB_HIGH LEVEL VALUE (H)" : Real = PLC TT426_5P_ALM_ANALOG_DB."HIGH LEVEL VALUE (H)" AT %DB2081.DBD30, 1 s
   "TT426_5P_ALM_ANALOG_DB_LOW LEVEL VALUE (L)" : Real = PLC TT426_5P_ALM_ANALOG_DB."LOW LEVEL VALUE (L)" AT %DB2081.DBD26, 1 s
   "TT426_5P_ALM_ANALOG_DB_VERY HIGH LEVEL VALUE (HH)" : Real = PLC TT426_5P_ALM_ANALOG_DB."VERY HIGH LEVEL VALUE (HH)" AT %DB2081.DBD34, 1 s
   "TT426_5P_ALM_ANALOG_DB_VERY LOW LEVEL VALUE (LL)" : Real = PLC TT426_5P_ALM_ANALOG_DB."VERY LOW LEVEL VALUE (LL)" AT %DB2081.DBD22, 1 s
   "TT426_5S_ALM_ANALOG_DB_HIGH LEVEL VALUE (H)" : Real = PLC TT426_5S_ALM_ANALOG_DB."HIGH LEVEL VALUE (H)" AT %DB2082.DBD30, 1 s
   "TT426_5S_ALM_ANALOG_DB_LOW LEVEL VALUE (L)" : Real = PLC TT426_5S_ALM_ANALOG_DB."LOW LEVEL VALUE (L)" AT %DB2082.DBD26, 1 s
